VERSION : 0.1
   VAR
      NewData : Bool := FALSE;
      FilteredShot : Array[1..10] of "UDT925_ShotResult";
      RealShot : Array[1..20] of "UDT925_ShotResult";
   END_VAR
BEGIN
   FilteredShot[1].PartNo := 0;
   FilteredShot[1].PartCounter := 0;
   FilteredShot[1].FoamingTime := 0.0;
   FilteredShot[1].PartWeight := 0.0;
   FilteredShot[1].StationNo := 16#00;
   FilteredShot[1].Machine_No := 16#00;
   FilteredShot[1].MHNo := 16#00;
   FilteredShot[1]."Name"[1] := '';
   FilteredShot[1]."Name"[2] := '';
   FilteredShot[1]."Name"[3] := '';
   FilteredShot[1]."Name"[4] := '';
   FilteredShot[1]."Name"[5] := '';
   FilteredShot[1]."Name"[6] := '';
   FilteredShot[1].Flow[1] := 0.0;
   FilteredShot[1].Flow[2] := 0.0;
   FilteredShot[1].Flow[3] := 0.0;
   FilteredShot[1].Flow[4] := 0.0;
   FilteredShot[1].Flow[5] := 0.0;
   FilteredShot[1].Flow[6] := 0.0;
   FilteredShot[1].Pressure[1] := 0.0;
   FilteredShot[1].Pressure[2] := 0.0;
   FilteredShot[1].Pressure[3] := 0.0;
   FilteredShot[1].Pressure[4] := 0.0;
   FilteredShot[1].Pressure[5] := 0.0;
   FilteredShot[1].Pressure[6] := 0.0;
   FilteredShot[1].Temperature[1] := 0.0;
   FilteredShot[1].Temperature[2] := 0.0;
   FilteredShot[1].Temperature[3] := 0.0;
   FilteredShot[1].Temperature[4] := 0.0;
   FilteredShot[1].Temperature[5] := 0.0;
   FilteredShot[1].Temperature[6] := 0.0;
   FilteredShot[1].MaterialConsumption[1] := 0.0;
   FilteredShot[1].MaterialConsumption[2] := 0.0;
   FilteredShot[1].MaterialConsumption[3] := 0.0;
   FilteredShot[1].MaterialConsumption[4] := 0.0;
   FilteredShot[1].MaterialConsumption[5] := 0.0;
   FilteredShot[1].MaterialConsumption[6] := 0.0;
   FilteredShot[1].Mixingratio[1] := 0.0;
   FilteredShot[1].Mixingratio[2] := 0.0;
   FilteredShot[1].Mixingratio[3] := 0.0;
   FilteredShot[1].Mixingratio[4] := 0.0;
   FilteredShot[1].Mixingratio[5] := 0.0;
   FilteredShot[1].Mixingratio[6] := 0.0;
   FilteredShot[1].StausBitWarning[1].StatusBitWarningMixingratio := FALSE;
   FilteredShot[1].StausBitWarning[1].StatusBitAlarmMixingratio := FALSE;
   FilteredShot[1].StausBitWarning[1].StatusBitWarningPressure := FALSE;
   FilteredShot[1].StausBitWarning[1].StatusBitAlarmPressure := FALSE;
   FilteredShot[1].StausBitWarning[1].StatusBitWarningPressureMH := FALSE;
   FilteredShot[1].StausBitWarning[1].StatusBitAlarmPressureMH := FALSE;
   FilteredShot[1].StausBitWarning[1].StatusBitWarningTemperature := FALSE;
   FilteredShot[1].StausBitWarning[1].StatusBitAlarmTemperature := FALSE;
   FilteredShot[1].StausBitWarning[1].StatusBitWarningTemperatureMH := FALSE;
   FilteredShot[1].StausBitWarning[1].StatusBitAlarmTemperatureMH := FALSE;
   FilteredShot[1].StausBitWarning[1].SpareBit11 := FALSE;
   FilteredShot[1].StausBitWarning[1].SpareBit12 := FALSE;
   FilteredShot[1].StausBitWarning[1].SpareBit13 := FALSE;
   FilteredShot[1].StausBitWarning[1].SpareBit14 := FALSE;
   FilteredShot[1].StausBitWarning[1].SpareBit15 := FALSE;
   FilteredShot[1].StausBitWarning[1].SpareBit16 := FALSE;
   FilteredShot[1].StausBitWarning[2].StatusBitWarningMixingratio := FALSE;
   FilteredShot[1].StausBitWarning[2].StatusBitAlarmMixingratio := FALSE;
   FilteredShot[1].StausBitWarning[2].StatusBitWarningPressure := FALSE;
   FilteredShot[1].StausBitWarning[2].StatusBitAlarmPressure := FALSE;
   FilteredShot[1].StausBitWarning[2].StatusBitWarningPressureMH := FALSE;
   FilteredShot[1].StausBitWarning[2].StatusBitAlarmPressureMH := FALSE;
   FilteredShot[1].StausBitWarning[2].StatusBitWarningTemperature := FALSE;
   FilteredShot[1].StausBitWarning[2].StatusBitAlarmTemperature := FALSE;
   FilteredShot[1].StausBitWarning[2].StatusBitWarningTemperatureMH := FALSE;
   FilteredShot[1].StausBitWarning[2].StatusBitAlarmTemperatureMH := FALSE;
   FilteredShot[1].StausBitWarning[2].SpareBit11 := FALSE;
   FilteredShot[1].StausBitWarning[2].SpareBit12 := FALSE;
   FilteredShot[1].StausBitWarning[2].SpareBit13 := FALSE;
   FilteredShot[1].StausBitWarning[2].SpareBit14 := FALSE;
   FilteredShot[1].StausBitWarning[2].SpareBit15 := FALSE;
   FilteredShot[1].StausBitWarning[2].SpareBit16 := FALSE;
   FilteredShot[1].StausBitWarning[3].StatusBitWarningMixingratio := FALSE;
   FilteredShot[1].StausBitWarning[3].StatusBitAlarmMixingratio := FALSE;
   FilteredShot[1].StausBitWarning[3].StatusBitWarningPressure := FALSE;
   FilteredShot[1].StausBitWarning[3].StatusBitAlarmPressure := FALSE;
   FilteredShot[1].StausBitWarning[3].StatusBitWarningPressureMH := FALSE;
   FilteredShot[1].StausBitWarning[3].StatusBitAlarmPressureMH := FALSE;
   FilteredShot[1].StausBitWarning[3].StatusBitWarningTemperature := FALSE;
   FilteredShot[1].StausBitWarning[3].StatusBitAlarmTemperature := FALSE;
   FilteredShot[1].StausBitWarning[3].StatusBitWarningTemperatureMH := FALSE;
   FilteredShot[1].StausBitWarning[3].StatusBitAlarmTemperatureMH := FALSE;
   FilteredShot[1].StausBitWarning[3].SpareBit11 := FALSE;
   FilteredShot[1].StausBitWarning[3].SpareBit12 := FALSE;
   FilteredShot[1].StausBitWarning[3].SpareBit13 := FALSE;
   FilteredShot[1].StausBitWarning[3].SpareBit14 := FALSE;
   FilteredShot[1].StausBitWarning[3].SpareBit15 := FALSE;
   FilteredShot[1].StausBitWarning[3].SpareBit16 := FALSE;
   FilteredShot[1].StausBitWarning[4].StatusBitWarningMixingratio := FALSE;
   FilteredShot[1].StausBitWarning[4].StatusBitAlarmMixingratio := FALSE;
   FilteredShot[1].StausBitWarning[4].StatusBitWarningPressure := FALSE;
   FilteredShot[1].StausBitWarning[4].StatusBitAlarmPressure := FALSE;
   FilteredShot[1].StausBitWarning[4].StatusBitWarningPressureMH := FALSE;
   FilteredShot[1].StausBitWarning[4].StatusBitAlarmPressureMH := FALSE;
   FilteredShot[1].StausBitWarning[4].StatusBitWarningTemperature := FALSE;
   FilteredShot[1].StausBitWarning[4].StatusBitAlarmTemperature := FALSE;
   FilteredShot[1].StausBitWarning[4].StatusBitWarningTemperatureMH := FALSE;
   FilteredShot[1].StausBitWarning[4].StatusBitAlarmTemperatureMH := FALSE;
   FilteredShot[1].StausBitWarning[4].SpareBit11 := FALSE;
   FilteredShot[1].StausBitWarning[4].SpareBit12 := FALSE;
   FilteredShot[1].StausBitWarning[4].SpareBit13 := FALSE;
   FilteredShot[1].StausBitWarning[4].SpareBit14 := FALSE;
   FilteredShot[1].StausBitWarning[4].SpareBit15 := FALSE;
   FilteredShot[1].StausBitWarning[4].SpareBit16 := FALSE;
   FilteredShot[1].StausBitWarning[5].StatusBitWarningMixingratio := FALSE;
   FilteredShot[1].StausBitWarning[5].StatusBitAlarmMixingratio := FALSE;
   FilteredShot[1].StausBitWarning[5].StatusBitWarningPressure := FALSE;
   FilteredShot[1].StausBitWarning[5].StatusBitAlarmPressure := FALSE;
   FilteredShot[1].StausBitWarning[5].StatusBitWarningPressureMH := FALSE;
   FilteredShot[1].StausBitWarning[5].StatusBitAlarmPressureMH := FALSE;
   FilteredShot[1].StausBitWarning[5].StatusBitWarningTemperature := FALSE;
   FilteredShot[1].StausBitWarning[5].StatusBitAlarmTemperature := FALSE;
   FilteredShot[1].StausBitWarning[5].StatusBitWarningTemperatureMH := FALSE;
   FilteredShot[1].StausBitWarning[5].StatusBitAlarmTemperatureMH := FALSE;
   FilteredShot[1].StausBitWarning[5].SpareBit11 := FALSE;
   FilteredShot[1].StausBitWarning[5].SpareBit12 := FALSE;
   FilteredShot[1].StausBitWarning[5].SpareBit13 := FALSE;
   FilteredShot[1].StausBitWarning[5].SpareBit14 := FALSE;
   FilteredShot[1].StausBitWarning[5].SpareBit15 := FALSE;
   FilteredShot[1].StausBitWarning[5].SpareBit16 := FALSE;
   FilteredShot[1].StausBitWarning[6].StatusBitWarningMixingratio := FALSE;
   FilteredShot[1].StausBitWarning[6].StatusBitAlarmMixingratio := FALSE;
   FilteredShot[1].StausBitWarning[6].StatusBitWarningPressure := FALSE;
   FilteredShot[1].StausBitWarning[6].StatusBitAlarmPressure := FALSE;
   FilteredShot[1].StausBitWarning[6].StatusBitWarningPressureMH := FALSE;
   FilteredShot[1].StausBitWarning[6].StatusBitAlarmPressureMH := FALSE;
   FilteredShot[1].StausBitWarning[6].StatusBitWarningTemperature := FALSE;
   FilteredShot[1].StausBitWarning[6].StatusBitAlarmTemperature := FALSE;
   FilteredShot[1].StausBitWarning[6].StatusBitWarningTemperatureMH := FALSE;
   FilteredShot[1].StausBitWarning[6].StatusBitAlarmTemperatureMH := FALSE;
   FilteredShot[1].StausBitWarning[6].SpareBit11 := FALSE;
   FilteredShot[1].StausBitWarning[6].SpareBit12 := FALSE;
   FilteredShot[1].StausBitWarning[6].SpareBit13 := FALSE;
   FilteredShot[1].StausBitWarning[6].SpareBit14 := FALSE;
   FilteredShot[1].StausBitWarning[6].SpareBit15 := FALSE;
   FilteredShot[1].StausBitWarning[6].SpareBit16 := FALSE;
   FilteredShot[1].PartShotDisableService := FALSE;
   FilteredShot[1].StatusBitFaultGroup1 := FALSE;
   FilteredShot[1].StatusBitStopCycleDuringShot := FALSE;
   FilteredShot[1].ShotDisabledDuringShot := FALSE;
   FilteredShot[1].StatusBitManualShot := FALSE;
   FilteredShot[1].StatusBitAutomaticShot := FALSE;
   FilteredShot[1].SpareBit7 := FALSE;
   FilteredShot[1].SpareBit8 := FALSE;
   FilteredShot[1].StatusBitWarningFlow := FALSE;
   FilteredShot[1].StatusBitAlarmFlow := FALSE;
   FilteredShot[1].StatusBitWarningWeight := FALSE;
   FilteredShot[1].StatusBitAlarmWeight := FALSE;
   FilteredShot[1].StatusBitWarningFoamingTime := FALSE;
   FilteredShot[1].StatusBitAlarmFoamingTime := FALSE;
   FilteredShot[1].SpareBit15 := FALSE;
   FilteredShot[1].SpareBit16 := FALSE;
   FilteredShot[2].PartNo := 0;
   FilteredShot[2].PartCounter := 0;
   FilteredShot[2].FoamingTime := 0.0;
   FilteredShot[2].PartWeight := 0.0;
   FilteredShot[2].StationNo := 16#00;
   FilteredShot[2].Machine_No := 16#00;
   FilteredShot[2].MHNo := 16#00;
   FilteredShot[2]."Name"[1] := '';
   FilteredShot[2]."Name"[2] := '';
   FilteredShot[2]."Name"[3] := '';
   FilteredShot[2]."Name"[4] := '';
   FilteredShot[2]."Name"[5] := '';
   FilteredShot[2]."Name"[6] := '';
   FilteredShot[2].Flow[1] := 0.0;
   FilteredShot[2].Flow[2] := 0.0;
   FilteredShot[2].Flow[3] := 0.0;
   FilteredShot[2].Flow[4] := 0.0;
   FilteredShot[2].Flow[5] := 0.0;
   FilteredShot[2].Flow[6] := 0.0;
   FilteredShot[2].Pressure[1] := 0.0;
   FilteredShot[2].Pressure[2] := 0.0;
   FilteredShot[2].Pressure[3] := 0.0;
   FilteredShot[2].Pressure[4] := 0.0;
   FilteredShot[2].Pressure[5] := 0.0;
   FilteredShot[2].Pressure[6] := 0.0;
   FilteredShot[2].Temperature[1] := 0.0;
   FilteredShot[2].Temperature[2] := 0.0;
   FilteredShot[2].Temperature[3] := 0.0;
   FilteredShot[2].Temperature[4] := 0.0;
   FilteredShot[2].Temperature[5] := 0.0;
   FilteredShot[2].Temperature[6] := 0.0;
   FilteredShot[2].MaterialConsumption[1] := 0.0;
   FilteredShot[2].MaterialConsumption[2] := 0.0;
   FilteredShot[2].MaterialConsumption[3] := 0.0;
   FilteredShot[2].MaterialConsumption[4] := 0.0;
   FilteredShot[2].MaterialConsumption[5] := 0.0;
   FilteredShot[2].MaterialConsumption[6] := 0.0;
   FilteredShot[2].Mixingratio[1] := 0.0;
   FilteredShot[2].Mixingratio[2] := 0.0;
   FilteredShot[2].Mixingratio[3] := 0.0;
   FilteredShot[2].Mixingratio[4] := 0.0;
   FilteredShot[2].Mixingratio[5] := 0.0;
   FilteredShot[2].Mixingratio[6] := 0.0;
   FilteredShot[2].StausBitWarning[1].StatusBitWarningMixingratio := FALSE;
   FilteredShot[2].StausBitWarning[1].StatusBitAlarmMixingratio := FALSE;
   // 4480 more start values not shown
END_DATA_BLOCK

DATA_BLOCK "DB919_ShotResultMach"   // DB919
TITLE = Shot result of last shot
{ S7_Optimized_Access := 'FALSE' }
VERSION : 0.1
   VAR
      ShotResult_Ma : Array[0..2] of "UDT919_ShotResult";
      TotalFlowShotM1 : Array[1..12] of Real;
      TotalFlowShotM2 : Array[1..12] of Real;
      AmountFlowValuesM1 : Array[1..12] of Real;
      AmountFlowValuesM2 : Array[1..12] of Real;
   END_VAR
BEGIN
END_DATA_BLOCK

DATA_BLOCK "DB925_ShotData_1"   // DB925
TITLE = Foaming: Shot set values RAM
{ S7_Optimized_Access := 'FALSE' }
AUTHOR : KT242
VERSION : 0.1
   VAR
      TimeStamp : DWord := 16#0000_0000;   // Time value of the last modification
      Shot_No_read : Int := 0;   // Number to write the shot to array[0]
      Shot_No_save : Int := 0;   // Number of shot to save at
      Shot_No_act : Word := 16#0000;   // Number of allcation at Shot[0]
      "Tool_No(1)" : Int := 0;   // Tool Number TEMP
      Tool_No : Int := 1;   // Tool Number
      Part_Shot_No : Int := 1;   // Part Shot Number
      Shots : Int := 0;
      Spare : Int := 0;
      CopyBit : Bool := FALSE;
      DataRead : Bool := FALSE;
      DataWrite : Bool := FALSE;
      "2PoinMovement_Comp01" : Bool := FALSE;
      "2PoinMovement_Comp02" : Bool := FALSE;
      "2PoinMovement_Comp03" : Bool := FALSE;
      "2PoinMovement_Comp04" : Bool := FALSE;
      "2PoinMovement_Comp05" : Bool := FALSE;
      "2PoinMovement_Comp06" : Bool := FALSE;
      Shot_TS1 : Int := 0;
      Shot_TS2 : Int := 0;
      Shot_TS3 : Int := 0;
      Shot_TS4 : Int := 0;
      Shot_TS5 : Int := 0;
      Shot_TS6 : Int := 0;
      Shot_TS7 : Int := 0;
      Shot_TS8 : Int := 0;
      Tool : Array[0.."AmountToolsDB"] of "UDT926_ShotSet";
   END_VAR
BEGIN
END_DATA_BLOCK

DATA_BLOCK "DB926_ShotData_2"   // DB926
TITLE = Foaming: Shot set values RAM
{ S7_Optimized_Access := 'FALSE' }
AUTHOR : KT242
VERSION : 0.1
   VAR
      Tool : Array[0.."AmountToolsDB"] of "UDT926_ShotSet";
   END_VAR
BEGIN
END_DATA_BLOCK

DATA_BLOCK "DB930_Tools"   // DB930
TITLE = Foaming: Tool values
{ S7_Optimized_Access := 'FALSE' }
VERSION : 0.1
   VAR
      TimeStamp : DWord := 16#0000_0000;
      Tool_No_read : Int := 0;
      Tool_No_save : Int := 0;
      Tool_No_act : Word := 16#0000;
      Tool : Array[0.."AmountTools"] of "UDT930_Tool";
      Delete_Impossible : Bool := FALSE;
   END_VAR
BEGIN
   Tool[0].Rob_Prog := 0;
   Tool[0].Rob_Prog2 := 0;
   Tool[0].PartShot_Amount := 16#01;
   Tool[0].EnableTool := TRUE;
   Tool[0].Spare5_2 := FALSE;
   Tool[0].Spare5_3 := FALSE;
   Tool[0].Spare5_4 := FALSE;
   Tool[0].Spare5_5 := FALSE;
   Tool[0].Spare5_6 := FALSE;
   Tool[0].EnablePurgeMH := FALSE;
   Tool[0].NitrogenVol := 0;
   Tool[0].Spare_12 := 16#0000;
   Tool[1].Rob_Prog := 0;
   Tool[1].Rob_Prog2 := 0;
   Tool[1].PartShot_Amount := 16#00;
   Tool[1].EnableTool := FALSE;
   Tool[1].Spare5_2 := FALSE;
   Tool[1].Spare5_3 := FALSE;
   Tool[1].Spare5_4 := FALSE;
   Tool[1].Spare5_5 := FALSE;
   Tool[1].Spare5_6 := FALSE;
   Tool[1].EnablePurgeMH := FALSE;
   Tool[1].NitrogenVol := 0;
   Tool[1].Spare_12 := 16#0000;
   Tool[2].Rob_Prog := 0;
   Tool[2].Rob_Prog2 := 0;
   Tool[2].PartShot_Amount := 16#00;
   Tool[2].EnableTool := FALSE;
   Tool[2].Spare5_2 := FALSE;
   Tool[2].Spare5_3 := FALSE;
   Tool[2].Spare5_4 := FALSE;
   Tool[2].Spare5_5 := FALSE;
   Tool[2].Spare5_6 := FALSE;
   Tool[2].EnablePurgeMH := FALSE;
   Tool[2].NitrogenVol := 0;
   Tool[2].Spare_12 := 16#0000;
   Tool[3].Rob_Prog := 0;
   Tool[3].Rob_Prog2 := 0;
   Tool[3].PartShot_Amount := 16#00;
   Tool[3].EnableTool := FALSE;
   Tool[3].Spare5_2 := FALSE;
   Tool[3].Spare5_3 := FALSE;
   Tool[3].Spare5_4 := FALSE;
   Tool[3].Spare5_5 := FALSE;
   Tool[3].Spare5_6 := FALSE;
   Tool[3].EnablePurgeMH := FALSE;
   Tool[3].NitrogenVol := 0;
   Tool[3].Spare_12 := 16#0000;
   Tool[4].Rob_Prog := 0;
   Tool[4].Rob_Prog2 := 0;
   Tool[4].PartShot_Amount := 16#00;
   Tool[4].EnableTool := FALSE;
   Tool[4].Spare5_2 := FALSE;
   Tool[4].Spare5_3 := FALSE;
   Tool[4].Spare5_4 := FALSE;
   Tool[4].Spare5_5 := FALSE;
   Tool[4].Spare5_6 := FALSE;
   Tool[4].EnablePurgeMH := FALSE;
   Tool[4].NitrogenVol := 0;
   Tool[4].Spare_12 := 16#0000;
   Tool[5].Rob_Prog := 0;
   Tool[5].Rob_Prog2 := 0;
   Tool[5].PartShot_Amount := 16#00;
   Tool[5].EnableTool := FALSE;
   Tool[5].Spare5_2 := FALSE;
   Tool[5].Spare5_3 := FALSE;
   Tool[5].Spare5_4 := FALSE;
   Tool[5].Spare5_5 := FALSE;
   Tool[5].Spare5_6 := FALSE;
   Tool[5].EnablePurgeMH := FALSE;
   Tool[5].NitrogenVol := 0;
   Tool[5].Spare_12 := 16#0000;
   Tool[6].Rob_Prog := 0;
   Tool[6].Rob_Prog2 := 0;
   Tool[6].PartShot_Amount := 16#00;
   Tool[6].EnableTool := FALSE;
   Tool[6].Spare5_2 := FALSE;
   Tool[6].Spare5_3 := FALSE;
   Tool[6].Spare5_4 := FALSE;
   Tool[6].Spare5_5 := FALSE;
   Tool[6].Spare5_6 := FALSE;
   Tool[6].EnablePurgeMH := FALSE;
   Tool[6].NitrogenVol := 0;
   Tool[6].Spare_12 := 16#0000;
   Tool[7].Rob_Prog := 0;
   Tool[7].Rob_Prog2 := 0;
   Tool[7].PartShot_Amount := 16#00;
   Tool[7].EnableTool := FALSE;
   Tool[7].Spare5_2 := FALSE;
   Tool[7].Spare5_3 := FALSE;
   Tool[7].Spare5_4 := FALSE;
   Tool[7].Spare5_5 := FALSE;
   Tool[7].Spare5_6 := FALSE;
   Tool[7].EnablePurgeMH := FALSE;
   Tool[7].NitrogenVol := 0;
   Tool[7].Spare_12 := 16#0000;
   Tool[8].Rob_Prog := 0;
   Tool[8].Rob_Prog2 := 0;
   Tool[8].PartShot_Amount := 16#00;
   Tool[8].EnableTool := FALSE;
   Tool[8].Spare5_2 := FALSE;
   Tool[8].Spare5_3 := FALSE;
   Tool[8].Spare5_4 := FALSE;
   Tool[8].Spare5_5 := FALSE;
   Tool[8].Spare5_6 := FALSE;
   Tool[8].EnablePurgeMH := FALSE;
   Tool[8].NitrogenVol := 0;
   Tool[8].Spare_12 := 16#0000;
   Tool[9].Rob_Prog := 0;
   Tool[9].Rob_Prog2 := 0;
   Tool[9].PartShot_Amount := 16#00;
   Tool[9].EnableTool := FALSE;
   Tool[9].Spare5_2 := FALSE;
   Tool[9].Spare5_3 := FALSE;
   Tool[9].Spare5_4 := FALSE;
   Tool[9].Spare5_5 := FALSE;
   Tool[9].Spare5_6 := FALSE;
   Tool[9].EnablePurgeMH := FALSE;
   Tool[9].NitrogenVol := 0;
   Tool[9].Spare_12 := 16#0000;
   Tool[10].Rob_Prog := 0;
   Tool[10].Rob_Prog2 := 0;
   Tool[10].PartShot_Amount := 16#00;
   Tool[10].EnableTool := FALSE;
   Tool[10].Spare5_2 := FALSE;
   Tool[10].Spare5_3 := FALSE;
   Tool[10].Spare5_4 := FALSE;
   Tool[10].Spare5_5 := FALSE;
   Tool[10].Spare5_6 := FALSE;
   Tool[10].EnablePurgeMH := FALSE;
   Tool[10].NitrogenVol := 0;
   Tool[10].Spare_12 := 16#0000;
   Tool[11].Rob_Prog := 0;
   Tool[11].Rob_Prog2 := 0;
   Tool[11].PartShot_Amount := 16#00;
   Tool[11].EnableTool := FALSE;
   Tool[11].Spare5_2 := FALSE;
   Tool[11].Spare5_3 := FALSE;
   Tool[11].Spare5_4 := FALSE;
   Tool[11].Spare5_5 := FALSE;
   Tool[11].Spare5_6 := FALSE;
   Tool[11].EnablePurgeMH := FALSE;
   Tool[11].NitrogenVol := 0;
   Tool[11].Spare_12 := 16#0000;
   Tool[12].Rob_Prog := 0;
   Tool[12].Rob_Prog2 := 0;
   Tool[12].PartShot_Amount := 16#00;
   Tool[12].EnableTool := FALSE;
   Tool[12].Spare5_2 := FALSE;
   Tool[12].Spare5_3 := FALSE;
   Tool[12].Spare5_4 := FALSE;
   Tool[12].Spare5_5 := FALSE;
   Tool[12].Spare5_6 := FALSE;
   Tool[12].EnablePurgeMH := FALSE;
   Tool[12].NitrogenVol := 0;
   Tool[12].Spare_12 := 16#0000;
   Tool[13].Rob_Prog := 0;
   Tool[13].Rob_Prog2 := 0;
   Tool[13].PartShot_Amount := 16#00;
   Tool[13].EnableTool := FALSE;
   Tool[13].Spare5_2 := FALSE;
   Tool[13].Spare5_3 := FALSE;
   Tool[13].Spare5_4 := FALSE;
   Tool[13].Spare5_5 := FALSE;
   Tool[13].Spare5_6 := FALSE;
   Tool[13].EnablePurgeMH := FALSE;
   Tool[13].NitrogenVol := 0;
   Tool[13].Spare_12 := 16#0000;
   Tool[14].Rob_Prog := 0;
   Tool[14].Rob_Prog2 := 0;
   Tool[14].PartShot_Amount := 16#00;
   Tool[14].EnableTool := FALSE;
   Tool[14].Spare5_2 := FALSE;
   Tool[14].Spare5_3 := FALSE;
   Tool[14].Spare5_4 := FALSE;
   Tool[14].Spare5_5 := FALSE;
   Tool[14].Spare5_6 := FALSE;
   Tool[14].EnablePurgeMH := FALSE;
   Tool[14].NitrogenVol := 0;
   Tool[14].Spare_12 := 16#0000;
   Tool[15].Rob_Prog := 0;
   Tool[15].Rob_Prog2 := 0;
   Tool[15].PartShot_Amount := 16#00;
   Tool[15].EnableTool := FALSE;
   Tool[15].Spare5_2 := FALSE;
   Tool[15].Spare5_3 := FALSE;
   Tool[15].Spare5_4 := FALSE;
   Tool[15].Spare5_5 := FALSE;
   Tool[15].Spare5_6 := FALSE;
   Tool[15].EnablePurgeMH := FALSE;
   Tool[15].NitrogenVol := 0;
   Tool[15].Spare_12 := 16#0000;
   Tool[16].Rob_Prog := 0;
   Tool[16].Rob_Prog2 := 0;
   Tool[16].PartShot_Amount := 16#00;
   Tool[16].EnableTool := FALSE;
   Tool[16].Spare5_2 := FALSE;
   Tool[16].Spare5_3 := FALSE;
   Tool[16].Spare5_4 := FALSE;
   Tool[16].Spare5_5 := FALSE;
   // 1214 more start values not shown
END_DATA_BLOCK

DATA_BLOCK "DB933_SaveSortProgs"   // DB933
TITLE = Sorted list of tools at machine
{ S7_Optimized_Access := 'FALSE' }
VERSION : 0.1
   VAR
      SaveSortTool : Array[0.."AmountTools"] of Int;
      ProgSort : Bool := FALSE;
   END_VAR
BEGIN
END_DATA_BLOCK

DATA_BLOCK "DB939_Tool_alloc_HMI"   // DB939
{ S7_Optimized_Access := 'TRUE' }
VERSION : 0.1
   VAR
      AllocList_page : Int;
      SavedProgs_page : Int;
      Selected_prog : Int;
      Selected_SavedProg : Int;   // Focus of the saved tools (usually 0)
      MH_No_selected : Int := 1;
      Limit_allocation_list : Int := 0;
      Limit_allocation_page : Int;
      Delete_selected_tool : Int;
      Operability_selected_line : Int;   // The programm number can be the tranfer to the alloc list by the operator
      Overwrite_selected_tool : Bool;   // overwrite the selected tool
      Overwrite_not_allowed : Bool;   // for PopUp
      "Delete_tool_in _all_allocations" : Bool;   // delete the selected tool in all allocation lists
      Tool_not_exist : Bool;   // for PopUp (not used)
      AllocList_decrease : Bool;
      AllocList_increase : Bool;
      SavedProgs_decrease : Bool;
      SavedProgs_increase : Bool;
      MH_Nr_decrease_visible : Bool;   // Bit for visibility of the arrows
      MH_Nr_increase_visible : Bool;   // Bit for visibility of the arrows
      AllocList_decrease_visible : Bool;   // Bit for visibility of the arrows
      AllocList_increase_visible : Bool;   // Bit for visibility of the arrows
      SavedProgs_decrease_visible : Bool;   // Bit for visibility of the arrows
      SavedProgs_increase_visible : Bool;   // Bit for visibility of the arrows
      Tool_allocation_automatic : Bool;
      Tool_allocation_manual : Bool;
      Select_hand_automatic_alloc : Bool;   // 0 - Automatic; 1 - Hand
      Alloc_stationTool : Array[0..30] of Int;
      Alloc_tool_name : Array[0..30] of String[20];
      SaveSortProgs : Array[0..20] of Int;
      SaveSortProg_name : Array[0..20] of String[20];
   END_VAR
BEGIN
   Alloc_stationTool[0] := 0;
   Alloc_stationTool[1] := 0;
   Alloc_stationTool[2] := 0;
   Alloc_stationTool[3] := 0;
   Alloc_stationTool[4] := 0;
   Alloc_stationTool[5] := 0;
   Alloc_stationTool[6] := 0;
   Alloc_stationTool[7] := 0;
   Alloc_stationTool[8] := 0;
   Alloc_stationTool[9] := 0;
   Alloc_stationTool[10] := 0;
   Alloc_stationTool[11] := 0;
   Alloc_stationTool[12] := 0;
   Alloc_stationTool[13] := 0;
   Alloc_stationTool[14] := 0;
   Alloc_stationTool[15] := 0;
   Alloc_stationTool[16] := 0;
   Alloc_stationTool[17] := 0;
   Alloc_stationTool[18] := 0;
   Alloc_stationTool[19] := 0;
   Alloc_stationTool[20] := 0;
   Alloc_stationTool[21] := 0;
   Alloc_stationTool[22] := 0;
   Alloc_stationTool[23] := 0;
   Alloc_stationTool[24] := 0;
   Alloc_stationTool[25] := 0;
   Alloc_stationTool[26] := 0;
   Alloc_stationTool[27] := 0;
   Alloc_stationTool[28] := 0;
   Alloc_stationTool[29] := 0;
   Alloc_stationTool[30] := 0;
END_DATA_BLOCK

DATA_BLOCK "DB940_Tool_alloc_automatic"   // DB940
{ S7_Optimized_Access := 'TRUE' }
VERSION : 0.1
   VAR RETAIN
      Alloc_stationTool : Array[0.."AmountAllocationAutomatic"] of Int;
   END_VAR
BEGIN
   Alloc_stationTool[0] := 0;
   Alloc_stationTool[1] := 0;
   Alloc_stationTool[2] := 0;
   Alloc_stationTool[3] := 0;
   Alloc_stationTool[4] := 0;
   Alloc_stationTool[5] := 0;
   Alloc_stationTool[6] := 0;
   Alloc_stationTool[7] := 0;
   Alloc_stationTool[8] := 0;
   Alloc_stationTool[9] := 0;
   Alloc_stationTool[10] := 0;
   Alloc_stationTool[11] := 0;
   Alloc_stationTool[12] := 0;
   Alloc_stationTool[13] := 0;
   Alloc_stationTool[14] := 0;
   Alloc_stationTool[15] := 0;
   Alloc_stationTool[16] := 0;
   Alloc_stationTool[17] := 0;
   Alloc_stationTool[18] := 0;
   Alloc_stationTool[19] := 0;
   Alloc_stationTool[20] := 0;
   Alloc_stationTool[21] := 0;
   Alloc_stationTool[22] := 0;
   Alloc_stationTool[23] := 0;
   Alloc_stationTool[24] := 0;
   Alloc_stationTool[25] := 0;
   Alloc_stationTool[26] := 0;
   Alloc_stationTool[27] := 0;
   Alloc_stationTool[28] := 0;
   Alloc_stationTool[29] := 0;
   Alloc_stationTool[30] := 0;
   Alloc_stationTool[31] := 0;
   Alloc_stationTool[32] := 0;
   Alloc_stationTool[33] := 0;
   Alloc_stationTool[34] := 0;
   Alloc_stationTool[35] := 0;
   Alloc_stationTool[36] := 0;
   Alloc_stationTool[37] := 0;
   Alloc_stationTool[38] := 0;
   Alloc_stationTool[39] := 0;
   Alloc_stationTool[40] := 0;
   Alloc_stationTool[41] := 0;
   Alloc_stationTool[42] := 0;
   Alloc_stationTool[43] := 0;
   Alloc_stationTool[44] := 0;
   Alloc_stationTool[45] := 0;
   Alloc_stationTool[46] := 0;
   Alloc_stationTool[47] := 0;
   Alloc_stationTool[48] := 0;
   Alloc_stationTool[49] := 0;
   Alloc_stationTool[50] := 0;
   Alloc_stationTool[51] := 0;
   Alloc_stationTool[52] := 0;
   Alloc_stationTool[53] := 0;
   Alloc_stationTool[54] := 0;
   Alloc_stationTool[55] := 0;
   Alloc_stationTool[56] := 0;
   Alloc_stationTool[57] := 0;
   Alloc_stationTool[58] := 0;
   Alloc_stationTool[59] := 0;
   Alloc_stationTool[60] := 0;
   Alloc_stationTool[61] := 0;
   Alloc_stationTool[62] := 0;
   Alloc_stationTool[63] := 0;
   Alloc_stationTool[64] := 0;
   Alloc_stationTool[65] := 0;
   Alloc_stationTool[66] := 0;
   Alloc_stationTool[67] := 0;
   Alloc_stationTool[68] := 0;
   Alloc_stationTool[69] := 0;
   Alloc_stationTool[70] := 0;
   Alloc_stationTool[71] := 0;
   Alloc_stationTool[72] := 0;
   Alloc_stationTool[73] := 0;
   Alloc_stationTool[74] := 0;
   Alloc_stationTool[75] := 0;
   Alloc_stationTool[76] := 0;
   Alloc_stationTool[77] := 0;
   Alloc_stationTool[78] := 0;
   Alloc_stationTool[79] := 0;
   Alloc_stationTool[80] := 0;
   Alloc_stationTool[81] := 0;
   Alloc_stationTool[82] := 0;
   Alloc_stationTool[83] := 0;
   Alloc_stationTool[84] := 0;
   Alloc_stationTool[85] := 0;
   Alloc_stationTool[86] := 0;
   Alloc_stationTool[87] := 0;
   Alloc_stationTool[88] := 0;
   Alloc_stationTool[89] := 0;
   Alloc_stationTool[90] := 0;
   Alloc_stationTool[91] := 0;
   Alloc_stationTool[92] := 0;
   Alloc_stationTool[93] := 0;
   Alloc_stationTool[94] := 0;
   Alloc_stationTool[95] := 0;
   Alloc_stationTool[96] := 0;
   Alloc_stationTool[97] := 0;
   Alloc_stationTool[98] := 0;
   Alloc_stationTool[99] := 0;
   Alloc_stationTool[100] := 0;
   Alloc_stationTool[101] := 0;
   Alloc_stationTool[102] := 0;
   Alloc_stationTool[103] := 0;
   Alloc_stationTool[104] := 0;
   Alloc_stationTool[105] := 0;
   Alloc_stationTool[106] := 0;
   Alloc_stationTool[107] := 0;
   Alloc_stationTool[108] := 0;
   Alloc_stationTool[109] := 0;
   Alloc_stationTool[110] := 0;
   Alloc_stationTool[111] := 0;
   Alloc_stationTool[112] := 0;
   Alloc_stationTool[113] := 0;
   Alloc_stationTool[114] := 0;
   Alloc_stationTool[115] := 0;
   Alloc_stationTool[116] := 0;
   Alloc_stationTool[117] := 0;
   Alloc_stationTool[118] := 0;
   Alloc_stationTool[119] := 0;
   Alloc_stationTool[120] := 0;
END_DATA_BLOCK

DATA_BLOCK "DB941_Tool_alloc_manual_MH"   // DB941
{ S7_Optimized_Access := 'TRUE' }
VERSION : 0.1
   VAR RETAIN
      MH : Array[1..16] of Struct
         Alloc_stationTool : Array[0..120] of Int;
      END_STRUCT;
   END_VAR
BEGIN
   MH[1].Alloc_stationTool[0] := 0;
   MH[1].Alloc_stationTool[1] := 0;
   MH[1].Alloc_stationTool[2] := 0;
   MH[1].Alloc_stationTool[3] := 0;
   MH[1].Alloc_stationTool[4] := 0;
   MH[1].Alloc_stationTool[5] := 0;
   MH[1].Alloc_stationTool[6] := 0;
   MH[1].Alloc_stationTool[7] := 0;
   MH[1].Alloc_stationTool[8] := 0;
   MH[1].Alloc_stationTool[9] := 0;
   MH[1].Alloc_stationTool[10] := 0;
   MH[1].Alloc_stationTool[11] := 0;
   MH[1].Alloc_stationTool[12] := 0;
   MH[1].Alloc_stationTool[13] := 0;
   MH[1].Alloc_stationTool[14] := 0;
   MH[1].Alloc_stationTool[15] := 0;
   MH[1].Alloc_stationTool[16] := 0;
   MH[1].Alloc_stationTool[17] := 0;
   MH[1].Alloc_stationTool[18] := 0;
   MH[1].Alloc_stationTool[19] := 0;
   MH[1].Alloc_stationTool[20] := 0;
   MH[1].Alloc_stationTool[21] := 0;
   MH[1].Alloc_stationTool[22] := 0;
   MH[1].Alloc_stationTool[23] := 0;
   MH[1].Alloc_stationTool[24] := 0;
   MH[1].Alloc_stationTool[25] := 0;
   MH[1].Alloc_stationTool[26] := 0;
   MH[1].Alloc_stationTool[27] := 0;
   MH[1].Alloc_stationTool[28] := 0;
   MH[1].Alloc_stationTool[29] := 0;
   MH[1].Alloc_stationTool[30] := 0;
   MH[1].Alloc_stationTool[31] := 0;
   MH[1].Alloc_stationTool[32] := 0;
   MH[1].Alloc_stationTool[33] := 0;
   MH[1].Alloc_stationTool[34] := 0;
   MH[1].Alloc_stationTool[35] := 0;
   MH[1].Alloc_stationTool[36] := 0;
   MH[1].Alloc_stationTool[37] := 0;
   MH[1].Alloc_stationTool[38] := 0;
   MH[1].Alloc_stationTool[39] := 0;
   MH[1].Alloc_stationTool[40] := 0;
   MH[1].Alloc_stationTool[41] := 0;
   MH[1].Alloc_stationTool[42] := 0;
   MH[1].Alloc_stationTool[43] := 0;
   MH[1].Alloc_stationTool[44] := 0;
   MH[1].Alloc_stationTool[45] := 0;
   MH[1].Alloc_stationTool[46] := 0;
   MH[1].Alloc_stationTool[47] := 0;
   MH[1].Alloc_stationTool[48] := 0;
   MH[1].Alloc_stationTool[49] := 0;
   MH[1].Alloc_stationTool[50] := 0;
   MH[1].Alloc_stationTool[51] := 0;
   MH[1].Alloc_stationTool[52] := 0;
   MH[1].Alloc_stationTool[53] := 0;
   MH[1].Alloc_stationTool[54] := 0;
   MH[1].Alloc_stationTool[55] := 0;
   MH[1].Alloc_stationTool[56] := 0;
   MH[1].Alloc_stationTool[57] := 0;
   MH[1].Alloc_stationTool[58] := 0;
   MH[1].Alloc_stationTool[59] := 0;
   MH[1].Alloc_stationTool[60] := 0;
   MH[1].Alloc_stationTool[61] := 0;
   MH[1].Alloc_stationTool[62] := 0;
   MH[1].Alloc_stationTool[63] := 0;
   MH[1].Alloc_stationTool[64] := 0;
   MH[1].Alloc_stationTool[65] := 0;
   MH[1].Alloc_stationTool[66] := 0;
   MH[1].Alloc_stationTool[67] := 0;
   MH[1].Alloc_stationTool[68] := 0;
   MH[1].Alloc_stationTool[69] := 0;
   MH[1].Alloc_stationTool[70] := 0;
   MH[1].Alloc_stationTool[71] := 0;
   MH[1].Alloc_stationTool[72] := 0;
   MH[1].Alloc_stationTool[73] := 0;
   MH[1].Alloc_stationTool[74] := 0;
   MH[1].Alloc_stationTool[75] := 0;
   MH[1].Alloc_stationTool[76] := 0;
   MH[1].Alloc_stationTool[77] := 0;
   MH[1].Alloc_stationTool[78] := 0;
   MH[1].Alloc_stationTool[79] := 0;
   MH[1].Alloc_stationTool[80] := 0;
   MH[1].Alloc_stationTool[81] := 0;
   MH[1].Alloc_stationTool[82] := 0;
   MH[1].Alloc_stationTool[83] := 0;
   MH[1].Alloc_stationTool[84] := 0;
   MH[1].Alloc_stationTool[85] := 0;
   MH[1].Alloc_stationTool[86] := 0;
   MH[1].Alloc_stationTool[87] := 0;
   MH[1].Alloc_stationTool[88] := 0;
   MH[1].Alloc_stationTool[89] := 0;
   MH[1].Alloc_stationTool[90] := 0;
   MH[1].Alloc_stationTool[91] := 0;
   MH[1].Alloc_stationTool[92] := 0;
   MH[1].Alloc_stationTool[93] := 0;
   MH[1].Alloc_stationTool[94] := 0;
   MH[1].Alloc_stationTool[95] := 0;
   MH[1].Alloc_stationTool[96] := 0;
   MH[1].Alloc_stationTool[97] := 0;
   MH[1].Alloc_stationTool[98] := 0;
   MH[1].Alloc_stationTool[99] := 0;
   MH[1].Alloc_stationTool[100] := 0;
END_DATA_BLOCK

DATA_BLOCK "DB1001_TT_State"   // DB1001
{ S7_Optimized_Access := 'FALSE' }
AUTHOR : KT242
VERSION : 0.1
   VAR
      Bits : Struct
         Taktdehnung : Bool;   // Es ist eine Taktzeitverlängerung angewählt
         Stop_fuer_WW : Bool;   // Die Anlage soll für einen Werkzeugwechsel gestoppt werden
         Stop_fuer_Teachen : Bool;   // Die Anlage soll für das Reinigen gestoppt werden
         StopAfterEmpty : Bool;   // Die Anlage soll stoppen nach dem Leerfahren
         Reserve_05 : Bool;
         Reserve_06 : Bool;
         Fault_Exist : Bool;   // A fault exist at the dryside
         Reserve_08 : Bool;
         Reserve_09 : Bool;
         CPCleaningLeftTurn : Bool;
         NoFoamingButton : Bool;
         TTEmptying : Bool;
         LastShotInTool : Bool;
         MHOpenForCleaning : Bool;
         Reserve_15 : Bool;
         Reserve_16 : Bool;
         Reserve_17 : Bool;
         Reserve_18 : Bool;
         Reserve_19 : Bool;
         Reserve_20 : Bool;
         Reserve_21 : Bool;
         Reserve_22 : Bool;
         Reserve_23 : Bool;
         Reserve_24 : Bool;
         Reserve_25 : Bool;
         Reserve_26 : Bool;
         Reserve_27 : Bool;
         Reserve_28 : Bool;
         Reserve_29 : Bool;
         Reserve_30 : Bool;
         Reserve_31 : Bool;
         Reserve_32 : Bool;
         Reserve_Word_04 : Word;
         Reserve_Word_06 : Word;
         Reserve_Word_08 : Word;
      END_STRUCT;
      BA_Anlage : "UDT_RT_Betriebsart";   // Status für die Betriebsart der Anlage
      Takt : "UDT_RT_Takt";   // Status für die Taktimpulsbildung der Anlage
      IPOS : "UDT_RT_IPOS";   // Status für die Ansteuerung des Antriebes der Anlage
      Segmentkennung : "UDT_RT_Station_Nr";   // Status für die Segment- und Positionsbildung der Anlage
      SegmentInfo : Array[1..32] of Struct
         Enable : Bool;
         ShotDone : Bool;
         Status : Int;
         SegmentNo : Int;
         FoamingProgram : Int;
      END_STRUCT;
      Kettenspanner : "UDT_RT_Kettenspanner";   // Status für die ANsteuerung des Kettenspanners
      Aktuelle_Position : Int;   // Die Aktuelle Position des Segmentes zur Referenzposition
      Segment_in_Position : Struct
         Reserve1 : Bool;
         Reserve6 : Bool;
         Start_Schaeumen : Bool;
         FRG_Schaeumen : Bool;
         Start_Trennen : Bool;
         Reserve2 : Bool;
         Reserve3 : Bool;
         Reserve4 : Bool;
         FRG_abloeschen_Programm : Bool;
         Reserve5 : Bool;
         Test_IFM_Initiator : Bool;
         Start_Bewegung_1 : Bool;
         Start_Bewegung_2 : Bool;
         Start_Bewegung_3 : Bool;
         Reserve_81_6 : Bool;
         Reserve_81_7 : Bool;
      END_STRUCT;
      SegmentReadyForFoaming : Array[1..32] of Bool;
      SegmentPreperationFoaming : Array[1..32] of Bool;
      SegmentEnableFoaming : Array[1..32] of Bool;
      SegmentShotEnds : Array[1..32] of Bool;
      SegmentWithFoam : Array[1..32] of Bool;
      SegmentToolExist : Array[1..32] of Bool;
      SegmentToolOpen : Array[1..32] of Bool;
      SegmentStatus : Array[1..32] of Int;
   END_VAR
BEGIN
END_DATA_BLOCK

DATA_BLOCK "PN_AI"   // DB1002
{ S7_Optimized_Access := 'FALSE' }
VERSION : 0.1
   VAR
      SetIndex : Int := 1;
      ActIndex : Int := 1;
      Send : Bool := FALSE;
      IndexError : Bool := FALSE;
      Module : Array[0..16] of Struct
         AI8 : "IDM_302_Analogin_Default_8";
         AIResistive_8 : "IDM_502_Analogin_Temperature_8";
         AO : Array[1..8] of "IDM_401_Analogout_Default";
      END_STRUCT;
   END_VAR
BEGIN
   Module[1].AI8.Address := 316;
   Module[1].AI8.X14_0.Data."Data[1]".Betriebsart := 16#02;
   Module[1].AIResistive_8.Address := 300;
   Module[1].AI8.X14_0.Data."Data[8]".Betriebsart := 16#02;
   Module[1].AI8.X14_0.Data."Data[7]".Betriebsart := 16#02;
   Module[1].AI8.X14_0.Data."Data[6]".Betriebsart := 16#02;
   Module[1].AI8.X14_0.Data."Data[5]".Betriebsart := 16#02;
   Module[1].AI8.X14_0.Data."Data[4]".Betriebsart := 16#02;
   Module[1].AI8.X14_0.Data."Data[3]".Betriebsart := 16#02;
   Module[1].AI8.X14_0.Data."Data[2]".Betriebsart := 16#02;
   Module[2].AI8.Address := 412;
   Module[2].AI8.X14_0.Data."Data[1]".Betriebsart := 16#02;
   Module[2].AI8.X14_0.Data."Data[8]".Betriebsart := 16#02;
   Module[2].AI8.X14_0.Data."Data[7]".Betriebsart := 16#02;
   Module[2].AI8.X14_0.Data."Data[6]".Betriebsart := 16#02;
   Module[2].AI8.X14_0.Data."Data[5]".Betriebsart := 16#02;
   Module[2].AI8.X14_0.Data."Data[4]".Betriebsart := 16#02;
   Module[2].AI8.X14_0.Data."Data[3]".Betriebsart := 16#02;
   Module[2].AI8.X14_0.Data."Data[2]".Betriebsart := 16#02;
   Module[2].AIResistive_8.Address := 396;
   Module[3].AI8.Address := 444;
   Module[3].AI8.X14_0.Data."Data[8]".Betriebsart := 16#02;
   Module[3].AI8.X14_0.Data."Data[7]".Betriebsart := 16#02;
   Module[3].AI8.X14_0.Data."Data[6]".Betriebsart := 16#02;
   Module[3].AI8.X14_0.Data."Data[5]".Betriebsart := 16#02;
   Module[3].AI8.X14_0.Data."Data[4]".Betriebsart := 16#02;
   Module[3].AI8.X14_0.Data."Data[3]".Betriebsart := 16#02;
   Module[3].AI8.X14_0.Data."Data[2]".Betriebsart := 16#02;
   Module[3].AI8.X14_0.Data."Data[1]".Betriebsart := 16#02;
   Module[3].AIResistive_8.Address := 428;
   Module[0].AI8.X14_0.Data."Data[1]".Betriebsart := 16#02;
   Module[0].AI8.X14_0.Data."Data[1]".Bereichsobergrenze := 6000;
   Module[0].AI8.X14_0.Data."Data[2]".Betriebsart := 16#02;
   Module[0].AI8.X14_0.Data."Data[2]".Bereichsobergrenze := 6000;
   Module[2].AI8.X14_0.Data."Data[2]".Bereichsobergrenze := 6000;
   Module[2].AI8.X14_0.Data."Data[1]".Bereichsobergrenze := 6000;
   Module[1].AI8.X14_0.Data."Data[2]".Bereichsobergrenze := 6000;
   Module[1].AI8.X14_0.Data."Data[1]".Bereichsobergrenze := 6000;
   Module[0].AI8.Address := 316;
   Module[0].AI8.Active := TRUE;
   Module[0].AI8.ChckConnFault := FALSE;
   Module[0].AI8.ChckConnDone := TRUE;
   Module[0].AI8.X14_0.Request := TRUE;
   Module[0].AI8.X14_0.Transmitting := TRUE;
   Module[0].AI8.X14_0.Active := FALSE;
   Module[0].AI8.X14_0.Data."Data[1]".Reserve := 16#00;
   Module[0].AI8.X14_0.Data."Data[1]".Bereichsuntergrenze := 0;
   Module[0].AI8.X14_0.Data."Data[1]".Mittelwertzeit := 200;
   Module[0].AI8.X14_0.Data."Data[2]".Reserve := 16#00;
   Module[0].AI8.X14_0.Data."Data[2]".Bereichsuntergrenze := 0;
   Module[0].AI8.X14_0.Data."Data[2]".Mittelwertzeit := 200;
   Module[0].AI8.X14_0.Data."Data[3]".Betriebsart := 16#02;
   Module[0].AI8.X14_0.Data."Data[3]".Reserve := 16#00;
   Module[0].AI8.X14_0.Data."Data[3]".Bereichsobergrenze := 1000;
   Module[0].AI8.X14_0.Data."Data[3]".Bereichsuntergrenze := 0;
   Module[0].AI8.X14_0.Data."Data[3]".Mittelwertzeit := 500;
   Module[0].AI8.X14_0.Data."Data[4]".Betriebsart := 16#02;
   Module[0].AI8.X14_0.Data."Data[4]".Reserve := 16#00;
   Module[0].AI8.X14_0.Data."Data[4]".Bereichsobergrenze := 1000;
   Module[0].AI8.X14_0.Data."Data[4]".Bereichsuntergrenze := 0;
   Module[0].AI8.X14_0.Data."Data[4]".Mittelwertzeit := 500;
   Module[0].AI8.X14_0.Data."Data[5]".Betriebsart := 16#02;
   Module[0].AI8.X14_0.Data."Data[5]".Reserve := 16#00;
   Module[0].AI8.X14_0.Data."Data[5]".Bereichsobergrenze := 1000;
   Module[0].AI8.X14_0.Data."Data[5]".Bereichsuntergrenze := 0;
   Module[0].AI8.X14_0.Data."Data[5]".Mittelwertzeit := 100;
   Module[0].AI8.X14_0.Data."Data[6]".Betriebsart := 16#02;
   Module[0].AI8.X14_0.Data."Data[6]".Reserve := 16#00;
   Module[0].AI8.X14_0.Data."Data[6]".Bereichsobergrenze := 1000;
   Module[0].AI8.X14_0.Data."Data[6]".Bereichsuntergrenze := 0;
   Module[0].AI8.X14_0.Data."Data[6]".Mittelwertzeit := 100;
   Module[0].AI8.X14_0.Data."Data[7]".Betriebsart := 16#02;
   Module[0].AI8.X14_0.Data."Data[7]".Reserve := 16#00;
   Module[0].AI8.X14_0.Data."Data[7]".Bereichsobergrenze := 1000;
   Module[0].AI8.X14_0.Data."Data[7]".Bereichsuntergrenze := 0;
   Module[0].AI8.X14_0.Data."Data[7]".Mittelwertzeit := 100;
   Module[0].AI8.X14_0.Data."Data[8]".Betriebsart := 16#02;
   Module[0].AI8.X14_0.Data."Data[8]".Reserve := 16#00;
   Module[0].AI8.X14_0.Data."Data[8]".Bereichsobergrenze := 6000;
   Module[0].AI8.X14_0.Data."Data[8]".Bereichsuntergrenze := 0;
   Module[0].AI8.X14_0.Data."Data[8]".Mittelwertzeit := 200;
   Module[0].AIResistive_8.Address := 300;
   Module[0].AIResistive_8.Active := TRUE;
   Module[0].AIResistive_8.ChckConnFault := FALSE;
   Module[0].AIResistive_8.ChckConnDone := TRUE;
   Module[0].AIResistive_8.TemperatureInput.Request := TRUE;
   Module[0].AIResistive_8.TemperatureInput.Transmitting := TRUE;
   Module[0].AIResistive_8.TemperatureInput.Active := FALSE;
   Module[0].AIResistive_8.TemperatureInput.Data[1].Mittelwertzeit := 100;
   Module[0].AIResistive_8.TemperatureInput.Data[1].ErsatzwertDrahtbruch := 0;
   Module[0].AIResistive_8.TemperatureInput.Data[1].Einheit := 16#00;
   Module[0].AIResistive_8.TemperatureInput.Data[1].Reserve := 16#00;
   Module[0].AIResistive_8.TemperatureInput.Data[2].Mittelwertzeit := 100;
   Module[0].AIResistive_8.TemperatureInput.Data[2].ErsatzwertDrahtbruch := 0;
   Module[0].AIResistive_8.TemperatureInput.Data[2].Einheit := 16#00;
   Module[0].AIResistive_8.TemperatureInput.Data[2].Reserve := 16#00;
   Module[0].AIResistive_8.TemperatureInput.Data[3].Mittelwertzeit := 100;
   Module[0].AIResistive_8.TemperatureInput.Data[3].ErsatzwertDrahtbruch := 0;
   Module[0].AIResistive_8.TemperatureInput.Data[3].Einheit := 16#00;
   Module[0].AIResistive_8.TemperatureInput.Data[3].Reserve := 16#00;
   Module[0].AIResistive_8.TemperatureInput.Data[4].Mittelwertzeit := 100;
   Module[0].AIResistive_8.TemperatureInput.Data[4].ErsatzwertDrahtbruch := 0;
   Module[0].AIResistive_8.TemperatureInput.Data[4].Einheit := 16#00;
   Module[0].AIResistive_8.TemperatureInput.Data[4].Reserve := 16#00;
   Module[0].AIResistive_8.TemperatureInput.Data[5].Mittelwertzeit := 100;
   Module[0].AIResistive_8.TemperatureInput.Data[5].ErsatzwertDrahtbruch := 0;
   Module[0].AIResistive_8.TemperatureInput.Data[5].Einheit := 16#00;
   Module[0].AIResistive_8.TemperatureInput.Data[5].Reserve := 16#00;
   Module[0].AIResistive_8.TemperatureInput.Data[6].Mittelwertzeit := 100;
   Module[0].AIResistive_8.TemperatureInput.Data[6].ErsatzwertDrahtbruch := 0;
   Module[0].AIResistive_8.TemperatureInput.Data[6].Einheit := 16#00;
   Module[0].AIResistive_8.TemperatureInput.Data[6].Reserve := 16#00;
   Module[0].AIResistive_8.TemperatureInput.Data[7].Mittelwertzeit := 100;
   Module[0].AIResistive_8.TemperatureInput.Data[7].ErsatzwertDrahtbruch := 0;
   Module[0].AIResistive_8.TemperatureInput.Data[7].Einheit := 16#00;
   Module[0].AIResistive_8.TemperatureInput.Data[7].Reserve := 16#00;
   Module[0].AIResistive_8.TemperatureInput.Data[8].Mittelwertzeit := 200;
   Module[0].AIResistive_8.TemperatureInput.Data[8].ErsatzwertDrahtbruch := 0;
   Module[0].AIResistive_8.TemperatureInput.Data[8].Einheit := 16#00;
   Module[0].AIResistive_8.TemperatureInput.Data[8].Reserve := 16#00;
   Module[0].AO[1].Address := 0;
   Module[0].AO[1].Active := FALSE;
   Module[0].AO[1].ChckConnFault := FALSE;
   Module[0].AO[1].ChckConnDone := FALSE;
   Module[0].AO[1].GeneralParameters.Request := FALSE;
   Module[0].AO[1].GeneralParameters.Transmitting := FALSE;
   Module[0].AO[1].GeneralParameters.Active := FALSE;
   Module[0].AO[1].GeneralParameters.Data.Ausgangskanal.Bit0 := FALSE;
   Module[0].AO[1].GeneralParameters.Data.Ausgangskanal.Bit1 := FALSE;
   Module[0].AO[1].GeneralParameters.Data.Ausgangskanal.Bit2 := FALSE;
   Module[0].AO[1].GeneralParameters.Data.Ausgangskanal.Spare3 := FALSE;
   Module[0].AO[1].GeneralParameters.Data.Ausgangskanal.Spare4 := FALSE;
   Module[0].AO[1].GeneralParameters.Data.Ausgangskanal.Spare5 := FALSE;
   Module[0].AO[1].GeneralParameters.Data.Ausgangskanal.Spare6 := FALSE;
   Module[0].AO[1].GeneralParameters.Data.Ausgangskanal.Spare7 := FALSE;
   Module[0].AO[1].GeneralParameters.Data.Ausgangskanal.Bereichsobergrenze := 10000;
   Module[0].AO[1].GeneralParameters.Data.Ausgangskanal.Bereichsuntergrenze := -10000;
   Module[0].AO[1].GeneralParameters.Data.Ausgangskanal.Rampenzeit := 1000;
   Module[0].AO[2].Address := 0;
   Module[0].AO[2].Active := FALSE;
   Module[0].AO[2].ChckConnFault := FALSE;
   Module[0].AO[2].ChckConnDone := FALSE;
   Module[0].AO[2].GeneralParameters.Request := FALSE;
   Module[0].AO[2].GeneralParameters.Transmitting := FALSE;
   Module[0].AO[2].GeneralParameters.Active := FALSE;
   Module[0].AO[2].GeneralParameters.Data.Ausgangskanal.Bit0 := FALSE;
   Module[0].AO[2].GeneralParameters.Data.Ausgangskanal.Bit1 := FALSE;
   Module[0].AO[2].GeneralParameters.Data.Ausgangskanal.Bit2 := FALSE;
   Module[0].AO[2].GeneralParameters.Data.Ausgangskanal.Spare3 := FALSE;
   Module[0].AO[2].GeneralParameters.Data.Ausgangskanal.Spare4 := FALSE;
   Module[0].AO[2].GeneralParameters.Data.Ausgangskanal.Spare5 := FALSE;
   Module[0].AO[2].GeneralParameters.Data.Ausgangskanal.Spare6 := FALSE;
   Module[0].AO[2].GeneralParameters.Data.Ausgangskanal.Spare7 := FALSE;
   Module[0].AO[2].GeneralParameters.Data.Ausgangskanal.Bereichsobergrenze := 10000;
   Module[0].AO[2].GeneralParameters.Data.Ausgangskanal.Bereichsuntergrenze := -10000;
   Module[0].AO[2].GeneralParameters.Data.Ausgangskanal.Rampenzeit := 1000;
   Module[0].AO[3].Address := 0;
   Module[0].AO[3].Active := FALSE;
   Module[0].AO[3].ChckConnFault := FALSE;
   Module[0].AO[3].ChckConnDone := FALSE;
   Module[0].AO[3].GeneralParameters.Request := FALSE;
   Module[0].AO[3].GeneralParameters.Transmitting := FALSE;
   Module[0].AO[3].GeneralParameters.Active := FALSE;
   Module[0].AO[3].GeneralParameters.Data.Ausgangskanal.Bit0 := FALSE;
   Module[0].AO[3].GeneralParameters.Data.Ausgangskanal.Bit1 := FALSE;
   Module[0].AO[3].GeneralParameters.Data.Ausgangskanal.Bit2 := FALSE;
   Module[0].AO[3].GeneralParameters.Data.Ausgangskanal.Spare3 := FALSE;
   Module[0].AO[3].GeneralParameters.Data.Ausgangskanal.Spare4 := FALSE;
   Module[0].AO[3].GeneralParameters.Data.Ausgangskanal.Spare5 := FALSE;
   Module[0].AO[3].GeneralParameters.Data.Ausgangskanal.Spare6 := FALSE;
   Module[0].AO[3].GeneralParameters.Data.Ausgangskanal.Spare7 := FALSE;
   Module[0].AO[3].GeneralParameters.Data.Ausgangskanal.Bereichsobergrenze := 10000;
   Module[0].AO[3].GeneralParameters.Data.Ausgangskanal.Bereichsuntergrenze := -10000;
   Module[0].AO[3].GeneralParameters.Data.Ausgangskanal.Rampenzeit := 1000;
   Module[0].AO[4].Address := 0;
   Module[0].AO[4].Active := FALSE;
   Module[0].AO[4].ChckConnFault := FALSE;
   Module[0].AO[4].ChckConnDone := FALSE;
   Module[0].AO[4].GeneralParameters.Request := FALSE;
   Module[0].AO[4].GeneralParameters.Transmitting := FALSE;
   Module[0].AO[4].GeneralParameters.Active := FALSE;
   Module[0].AO[4].GeneralParameters.Data.Ausgangskanal.Bit0 := FALSE;
   Module[0].AO[4].GeneralParameters.Data.Ausgangskanal.Bit1 := FALSE;
   Module[0].AO[4].GeneralParameters.Data.Ausgangskanal.Bit2 := FALSE;
   Module[0].AO[4].GeneralParameters.Data.Ausgangskanal.Spare3 := FALSE;
   Module[0].AO[4].GeneralParameters.Data.Ausgangskanal.Spare4 := FALSE;
   Module[0].AO[4].GeneralParameters.Data.Ausgangskanal.Spare5 := FALSE;
   Module[0].AO[4].GeneralParameters.Data.Ausgangskanal.Spare6 := FALSE;
   Module[0].AO[4].GeneralParameters.Data.Ausgangskanal.Spare7 := FALSE;
   Module[0].AO[4].GeneralParameters.Data.Ausgangskanal.Bereichsobergrenze := 10000;
   Module[0].AO[4].GeneralParameters.Data.Ausgangskanal.Bereichsuntergrenze := -10000;
   Module[0].AO[4].GeneralParameters.Data.Ausgangskanal.Rampenzeit := 1000;
   Module[0].AO[5].Address := 0;
   Module[0].AO[5].Active := FALSE;
   Module[0].AO[5].ChckConnFault := FALSE;
   Module[0].AO[5].ChckConnDone := FALSE;
   Module[0].AO[5].GeneralParameters.Request := FALSE;
   Module[0].AO[5].GeneralParameters.Transmitting := FALSE;
   Module[0].AO[5].GeneralParameters.Active := FALSE;
   Module[0].AO[5].GeneralParameters.Data.Ausgangskanal.Bit0 := FALSE;
   // 3710 more start values not shown
END_DATA_BLOCK

